(* Logix 5000 project; controller MV vendor 1 type 14 code 217 rev 31.11; software revision 31.00; part 14 of 53 *)
(* tags used below, declared in another part *)
   CWD : CHECKWORD_FLAGS;
   MC_copy_how_many : DINT;
   MC_data_file_value_to_move : DINT;
   MC_Delphi_I : DINT[60];
   MC_from_data_file : DINT;
   MC_from_data_offset : DINT;
   MC_LTX_001_1 : PlantItem;   // LTX_001_1
   MC_LTX_001_2 : PlantItem;   // LTX_001_2
   MC_LTX_001_3 : PlantItem;   // LTX_001_3
   MC_LTX_002_1 : PlantItem;   // LTX_002_1
   MC_LTX_002_2 : PlantItem;   // LTX_002_2
   MC_LTX_002_3 : PlantItem;   // LTX_002_3
   MC_LTX_003_1 : PlantItem;   // LTX_003_1
   MC_LTX_003_2 : PlantItem;   // LTX_003_2
   MC_LTX_003_3 : PlantItem;   // LTX_003_3
   MC_N10 : INT[255];   // SETTINGS
   MC_N100 : INT[255];   // C1_PLC Channel 1 PLC data
   MC_N101 : INT[255];   // CH1 PC>PLC Channel 1 PC to PLC
   MC_N102 : INT[255];   // CH1 PROG Channel 1 CIP progra m
   MC_N103 : INT[255];   // CH1 ITEMS Chwd.nos.of items to be checked for Chan nel 1
   MC_N104 : INT[255];   // CH1 REPORT Channel 1 CIP report file
   MC_N108 : INT[255];   // CH1 VDATA Channel 1 CIP progra m validation data
   MC_N112 : INT[255];   // FVR DATA Data read from FV ro uting PLC
   MC_N113 : INT[255];   // MVR DATA Data read from MV ro uting PLC
   MC_N114 : INT[255];   // YP DATA
   MC_N120 : INT[255];   // C2 PLC Channel 2 PLC data
   MC_N121 : INT[255];   // CH2 PC>PLC Channel 2 PC to PLC
   MC_N122 : INT[255];   // CH2 PROG Channel 2 CIP progra m
   MC_N123 : INT[255];   // CH2 ITEMS Chwd.nos.of items to be checked for Chan nel 2
   MC_N124 : INT[255];   // CH2 REPORT Channel 2 CIP report file
   MC_N128 : INT[255];   // CH2 VDATA Channel 2 CIP progra m validation data
   MC_N160 : INT[255];   // P40 CHECK
   MC_N161 : INT[255];   // P41 CHECK
   MC_N162 : INT[255];   // P42 CHECK
   MC_N163 : INT[255];   // P43 CHECK
   MC_N164 : INT[255];   // P44 CHECK
   MC_N165 : INT[255];   // P45 CHECK
   MC_N166 : INT[255];   // P46 CHECK
   MC_N167 : INT[255];   // Original N File From SLC, No Description Available
   MC_N20 : INT[255];   // P1 PRESS Control block and da ta for P1 pressure P ID loop
   MC_N200 : INT[255];   // CHK_WORK Plant item fault che cking work area
   MC_N201 : INT[255];   // P1 CHECK CIP program 1 plant item check list
   MC_N202 : INT[255];   // P2 CHECK CIP program 2 plant item check list
   MC_N203 : INT[255];   // P3 CHECK CIP program 3 plant item check list
   MC_N204 : INT[255];   // P4 CHECK CIP program 4 plant item check list
   MC_N205 : INT[255];   // P5 CHECK CIP program 5 plant item check list
   MC_N206 : INT[255];   // P6 CHECK CIP program 6 plant item check list
   MC_N207 : INT[255];   // P7 CHECK CIP program 7 plant item check list
   MC_N208 : INT[255];   // P8 CHECK CIP program 8 plant item check list
   MC_N209 : INT[255];   // P9 CHECK CIP program 9 plant item check list
   MC_N21 : INT[255];   // P1 FLOW Control block and da ta for P1 flowrate P ID loop
   MC_N210 : INT[255];   // P10 CHECK CIP program 10 plant item check list
   MC_N211 : INT[255];   // P11 CHECK CIP program 11 plant item check list
   MC_N212 : INT[255];   // P12 CHECK CIP program 12 plant item check list
   MC_N213 : INT[255];   // P13 CHECK CIP program 13 plant item check list
   MC_N214 : INT[255];   // P14 CHECK CIP program 14 plant item check list
   MC_N215 : INT[255];   // P15 CHECK CIP program 15 plant item check list
   MC_N216 : INT[255];   // P16 CHECK CIP program 16 plant item check list
   MC_N217 : INT[255];   // P17 CHECK CIP program 17 plant item check list
   MC_N218 : INT[255];   // P18 CHECK CIP program 18 plant item check list
   MC_N219 : INT[255];   // P19 CHECK CIP program 19 plant item check list
   MC_N22 : INT[255];   // P2 PRESS Control block and da ta for P2 pressure P ID loop
   MC_N220 : INT[255];   // P20 CHECK CIP program 20 plant item check list
   MC_N221 : INT[255];   // P21 CHECK CIP program 21 plant item check list
   MC_N222 : INT[255];   // P22 CHECK CIP program 22 plant item check list
   MC_N223 : INT[255];   // P23 CHECK CIP program 23 plant item check list
   MC_N224 : INT[255];   // P24 CHECK CIP program 24 plant item check list
   MC_N225 : INT[255];   // P25 CHECK CIP program 25 plant item check list
   MC_N226 : INT[255];   // P26 CHECK CIP program 26 plant item check list
   MC_N227 : INT[255];   // P27 CHECK CIP program 27 plant item check list
   MC_N228 : INT[255];   // P28 CHECK CIP program 28 plant item check list
   MC_N229 : INT[255];   // P29 CHECK CIP program 29 plant item check list
   MC_N23 : INT[255];   // P2 FLOW Control block and da ta for P2 flowrate P ID loop
   MC_N230 : INT[255];   // P30 CHECK CIP program 30 plant item check list
   MC_N231 : INT[255];   // P31 CHECK CIP program 31 plant item check list
   MC_N232 : INT[255];   // P32 CHECK CIP program 32 plant item check list
   MC_N233 : INT[255];   // P33 CHECK CIP program 33 plant item check list
   MC_N234 : INT[255];   // P34 CHECK CIP program 34 plant item check list
   MC_N235 : INT[255];   // P35 CHECK CIP program 35 plant item check list
   MC_N236 : INT[255];   // P36 CHECK CIP program 36 plant item check list
   MC_N237 : INT[255];   // P37 CHECK CIP program 37 plant item check list
   MC_N238 : INT[255];   // P38 CHECK CIP program 38 plant item check list
   MC_N239 : INT[255];   // P39 CHECK CIP program 39 plant item check list
   MC_N245 : INT[255];   // CC_WORK Continuous checking program work area
   MC_N7 : INT[255];   // INTEGER
   MC_N80 : INT[255];   // SRV1_PLC Detergent tank 1 ser vice PLC data
   MC_N81 : INT[255];   // SV1_PC Detergent tank 1 ser vice PC to PLC data
   MC_N82 : INT[255];   // SV1 ITEMS Chwd.nos.of items to be checked for DT1 service
   MC_N90 : INT[255];   // SV2_PLC Detergent tank 2 ser vice PLC data
   MC_N91 : INT[255];   // SV2_PC Detergent tank 2 ser vice PC to PLC data
   MC_N92 : INT[255];   // SV2 ITEMS Chwd.nos.of items to be checked for DT2 service
   MC_PX_100 : PlantItem;   // PX_100
   MC_PX_100_RawInput : ALIAS FOR RIO_Rack_2:11:I.Data.18;   // MC_PX_100
   MC_PX_101 : PlantItem;   // PX_101
   MC_PX_101_RawInput : ALIAS FOR RIO_Rack_2:11:I.Data.19;   // MC_PX_101
   MC_R2_SW1 : PlantItem;   // R2_SW1
   MC_R2_SW1_RawInput : ALIAS FOR RIO_Rack_2:12:I.Data.0;   // MC_R2_SW1
   MC_R2_SW2 : PlantItem;   // R2_SW2
   MC_R2_SW2_RawInput : ALIAS FOR RIO_Rack_2:12:I.Data.1;   // MC_R2_SW2
   MC_R2_SW3 : PlantItem;   // R2_SW3
   MC_R2_SW3_1 : PlantItem;   // R2_SW3_1
   MC_R2_SW3_1_RawInput : ALIAS FOR RIO_Rack_2:12:I.Data.3;   // MC_R2_SW3_1
   MC_R2_SW3_RawInput : ALIAS FOR RIO_Rack_2:12:I.Data.2;   // MC_R2_SW3
   MC_R2_SW4 : PlantItem;   // R2_SW4
   MC_R2_SW4_RawInput : ALIAS FOR RIO_Rack_2:12:I.Data.4;   // MC_R2_SW4
   MC_R3_SW1 : PlantItem;   // R3_SW1
   MC_R3_SW1_RawInput : ALIAS FOR RIO_Rack_2:12:I.Data.5;   // MC_R3_SW1
   MC_R3_SW2 : PlantItem;   // R3_SW2
   MC_R3_SW2_RawInput : ALIAS FOR RIO_Rack_2:12:I.Data.6;   // MC_R3_SW2
   MC_T4 : TIMER[255];   // TIMER
   MC_to_data_file : DINT;
   MC_to_data_offset : DINT;
   One_Second_One_Scan : ALIAS FOR One_Second_1_scan;
(* MC_Common, continued *)

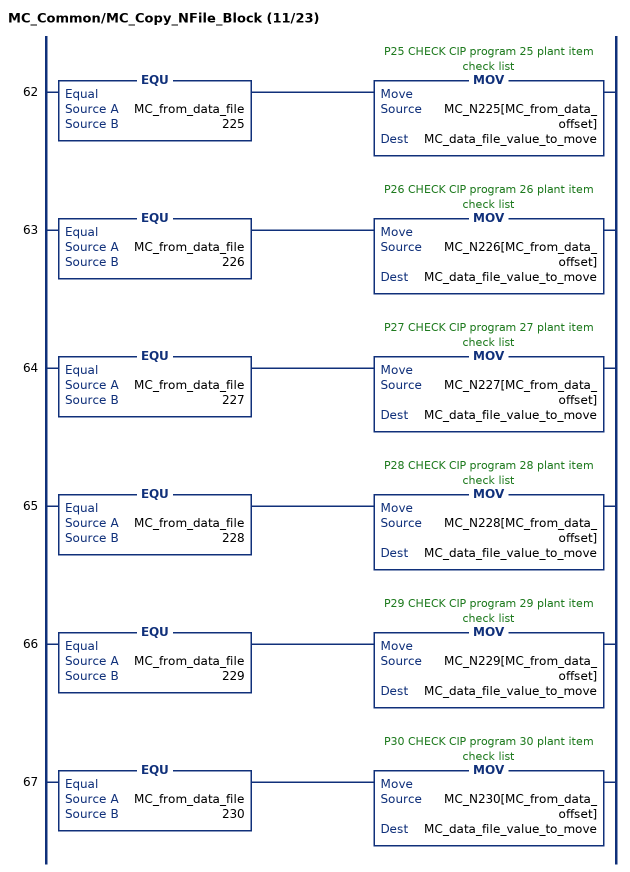
   [picture p203: MC_Common/MC_Copy_NFile_Block rungs 62-67]
   62: EQU(MC_from_data_file,225)MOV(MC_N225[MC_from_data_offset],MC_data_file_value_to_move);
   63: EQU(MC_from_data_file,226)MOV(MC_N226[MC_from_data_offset],MC_data_file_value_to_move);
   64: EQU(MC_from_data_file,227)MOV(MC_N227[MC_from_data_offset],MC_data_file_value_to_move);
   65: EQU(MC_from_data_file,228)MOV(MC_N228[MC_from_data_offset],MC_data_file_value_to_move);
   66: EQU(MC_from_data_file,229)MOV(MC_N229[MC_from_data_offset],MC_data_file_value_to_move);
   67: EQU(MC_from_data_file,230)MOV(MC_N230[MC_from_data_offset],MC_data_file_value_to_move);
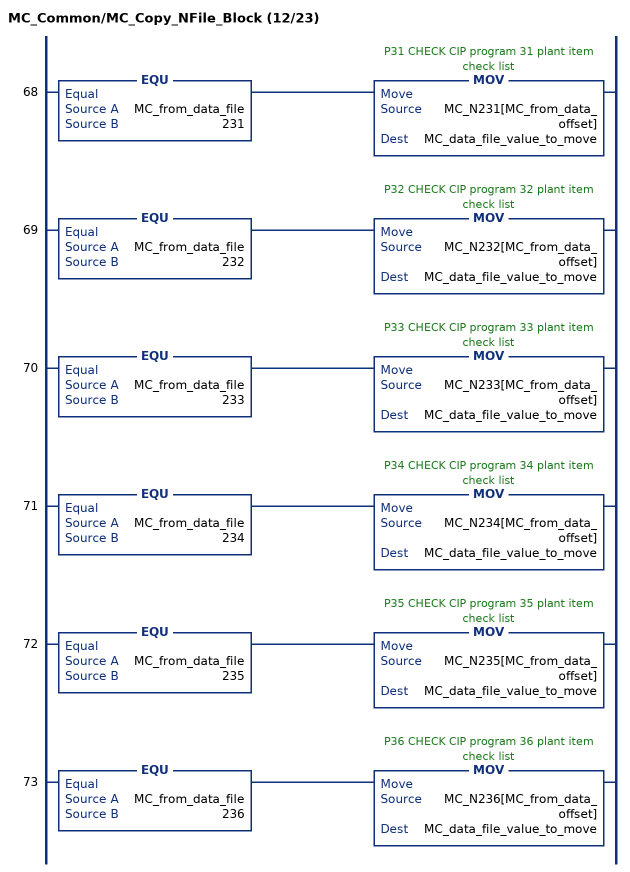
   68: EQU(MC_from_data_file,231)MOV(MC_N231[MC_from_data_offset],MC_data_file_value_to_move);
   69: EQU(MC_from_data_file,232)MOV(MC_N232[MC_from_data_offset],MC_data_file_value_to_move);
   70: EQU(MC_from_data_file,233)MOV(MC_N233[MC_from_data_offset],MC_data_file_value_to_move);
   71: EQU(MC_from_data_file,234)MOV(MC_N234[MC_from_data_offset],MC_data_file_value_to_move);
   72: EQU(MC_from_data_file,235)MOV(MC_N235[MC_from_data_offset],MC_data_file_value_to_move);
   73: EQU(MC_from_data_file,236)MOV(MC_N236[MC_from_data_offset],MC_data_file_value_to_move);
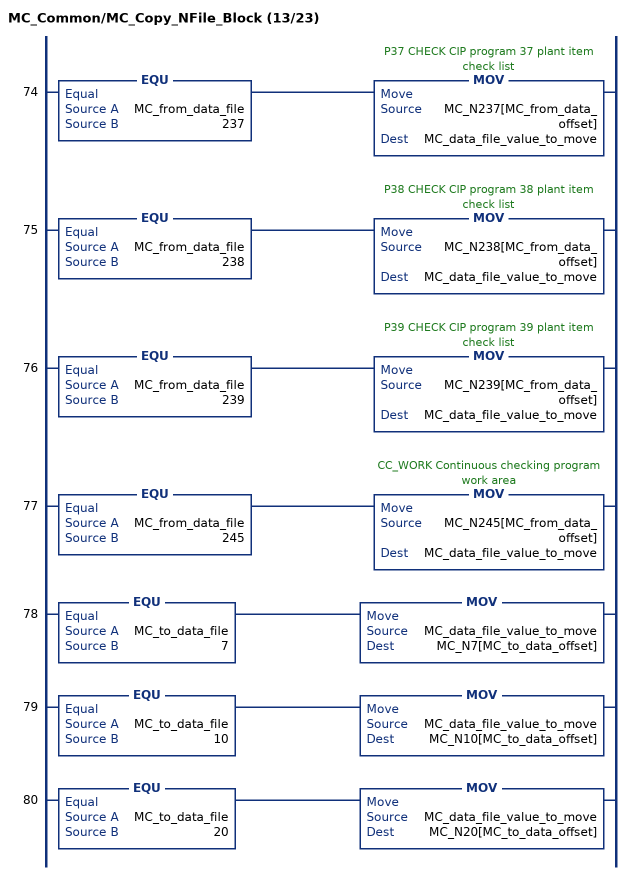
   74: EQU(MC_from_data_file,237)MOV(MC_N237[MC_from_data_offset],MC_data_file_value_to_move);
   75: EQU(MC_from_data_file,238)MOV(MC_N238[MC_from_data_offset],MC_data_file_value_to_move);
   76: EQU(MC_from_data_file,239)MOV(MC_N239[MC_from_data_offset],MC_data_file_value_to_move);
   77: EQU(MC_from_data_file,245)MOV(MC_N245[MC_from_data_offset],MC_data_file_value_to_move);
   78: EQU(MC_to_data_file,7)MOV(MC_data_file_value_to_move,MC_N7[MC_to_data_offset]);
   79: EQU(MC_to_data_file,10)MOV(MC_data_file_value_to_move,MC_N10[MC_to_data_offset]);
   80: EQU(MC_to_data_file,20)MOV(MC_data_file_value_to_move,MC_N20[MC_to_data_offset]);
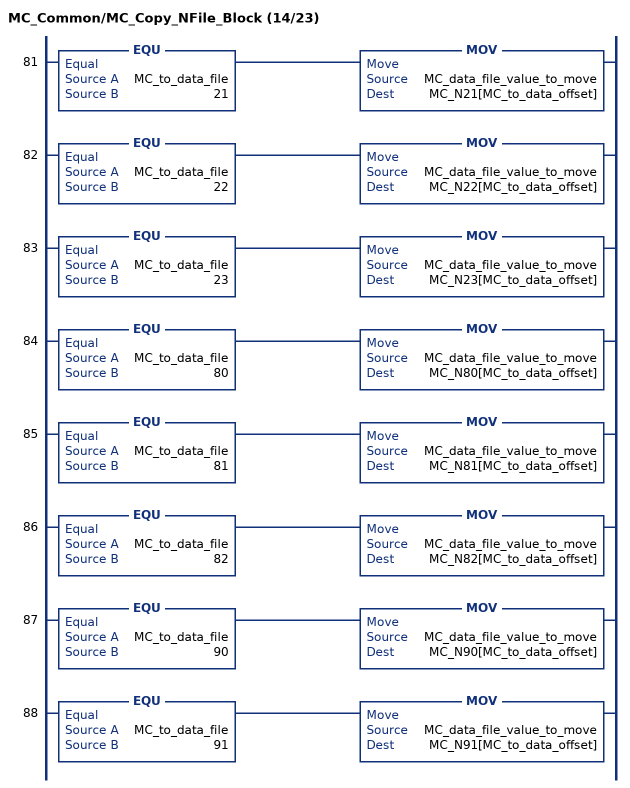
   81: EQU(MC_to_data_file,21)MOV(MC_data_file_value_to_move,MC_N21[MC_to_data_offset]);
   82: EQU(MC_to_data_file,22)MOV(MC_data_file_value_to_move,MC_N22[MC_to_data_offset]);
   83: EQU(MC_to_data_file,23)MOV(MC_data_file_value_to_move,MC_N23[MC_to_data_offset]);
   84: EQU(MC_to_data_file,80)MOV(MC_data_file_value_to_move,MC_N80[MC_to_data_offset]);
   85: EQU(MC_to_data_file,81)MOV(MC_data_file_value_to_move,MC_N81[MC_to_data_offset]);
   86: EQU(MC_to_data_file,82)MOV(MC_data_file_value_to_move,MC_N82[MC_to_data_offset]);
   87: EQU(MC_to_data_file,90)MOV(MC_data_file_value_to_move,MC_N90[MC_to_data_offset]);
   88: EQU(MC_to_data_file,91)MOV(MC_data_file_value_to_move,MC_N91[MC_to_data_offset]);
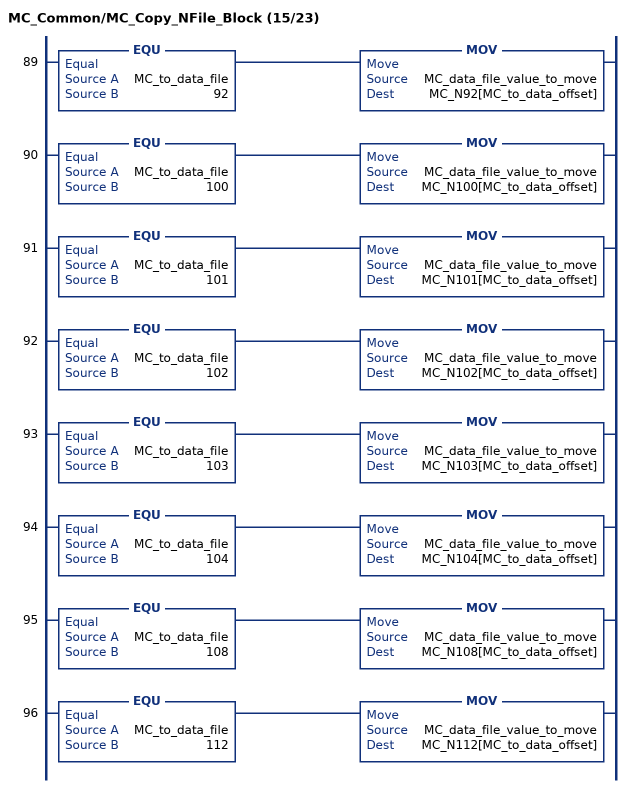
   89: EQU(MC_to_data_file,92)MOV(MC_data_file_value_to_move,MC_N92[MC_to_data_offset]);
   90: EQU(MC_to_data_file,100)MOV(MC_data_file_value_to_move,MC_N100[MC_to_data_offset]);
   91: EQU(MC_to_data_file,101)MOV(MC_data_file_value_to_move,MC_N101[MC_to_data_offset]);
   92: EQU(MC_to_data_file,102)MOV(MC_data_file_value_to_move,MC_N102[MC_to_data_offset]);
   93: EQU(MC_to_data_file,103)MOV(MC_data_file_value_to_move,MC_N103[MC_to_data_offset]);
   94: EQU(MC_to_data_file,104)MOV(MC_data_file_value_to_move,MC_N104[MC_to_data_offset]);
   95: EQU(MC_to_data_file,108)MOV(MC_data_file_value_to_move,MC_N108[MC_to_data_offset]);
   96: EQU(MC_to_data_file,112)MOV(MC_data_file_value_to_move,MC_N112[MC_to_data_offset]);
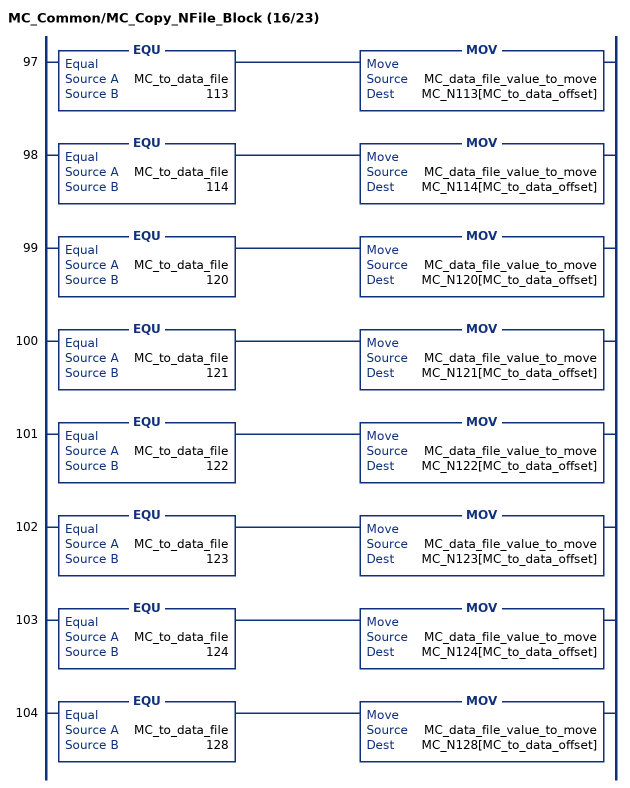
   97: EQU(MC_to_data_file,113)MOV(MC_data_file_value_to_move,MC_N113[MC_to_data_offset]);
   98: EQU(MC_to_data_file,114)MOV(MC_data_file_value_to_move,MC_N114[MC_to_data_offset]);
   99: EQU(MC_to_data_file,120)MOV(MC_data_file_value_to_move,MC_N120[MC_to_data_offset]);
   100: EQU(MC_to_data_file,121)MOV(MC_data_file_value_to_move,MC_N121[MC_to_data_offset]);
   101: EQU(MC_to_data_file,122)MOV(MC_data_file_value_to_move,MC_N122[MC_to_data_offset]);
   102: EQU(MC_to_data_file,123)MOV(MC_data_file_value_to_move,MC_N123[MC_to_data_offset]);
   103: EQU(MC_to_data_file,124)MOV(MC_data_file_value_to_move,MC_N124[MC_to_data_offset]);
   104: EQU(MC_to_data_file,128)MOV(MC_data_file_value_to_move,MC_N128[MC_to_data_offset]);
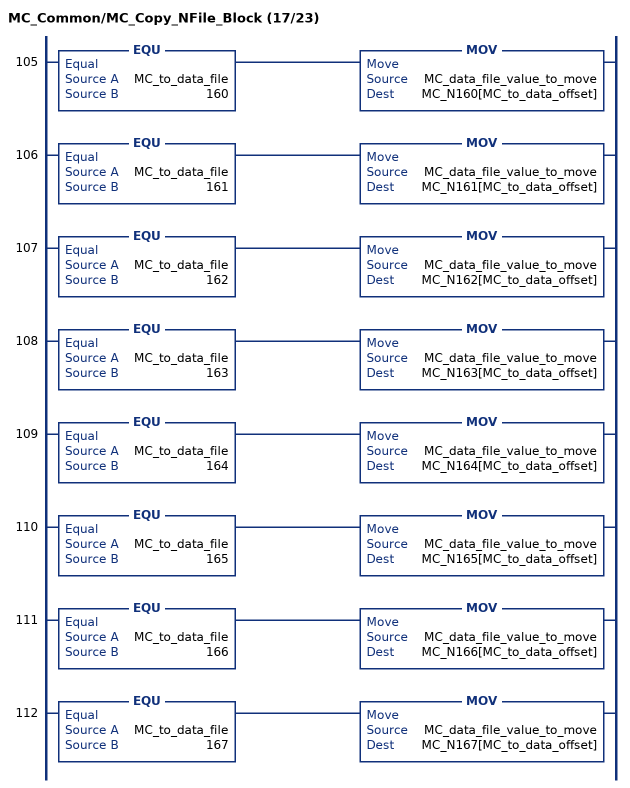
   105: EQU(MC_to_data_file,160)MOV(MC_data_file_value_to_move,MC_N160[MC_to_data_offset]);
   106: EQU(MC_to_data_file,161)MOV(MC_data_file_value_to_move,MC_N161[MC_to_data_offset]);
   107: EQU(MC_to_data_file,162)MOV(MC_data_file_value_to_move,MC_N162[MC_to_data_offset]);
   108: EQU(MC_to_data_file,163)MOV(MC_data_file_value_to_move,MC_N163[MC_to_data_offset]);
   109: EQU(MC_to_data_file,164)MOV(MC_data_file_value_to_move,MC_N164[MC_to_data_offset]);
   110: EQU(MC_to_data_file,165)MOV(MC_data_file_value_to_move,MC_N165[MC_to_data_offset]);
   111: EQU(MC_to_data_file,166)MOV(MC_data_file_value_to_move,MC_N166[MC_to_data_offset]);
   112: EQU(MC_to_data_file,167)MOV(MC_data_file_value_to_move,MC_N167[MC_to_data_offset]);
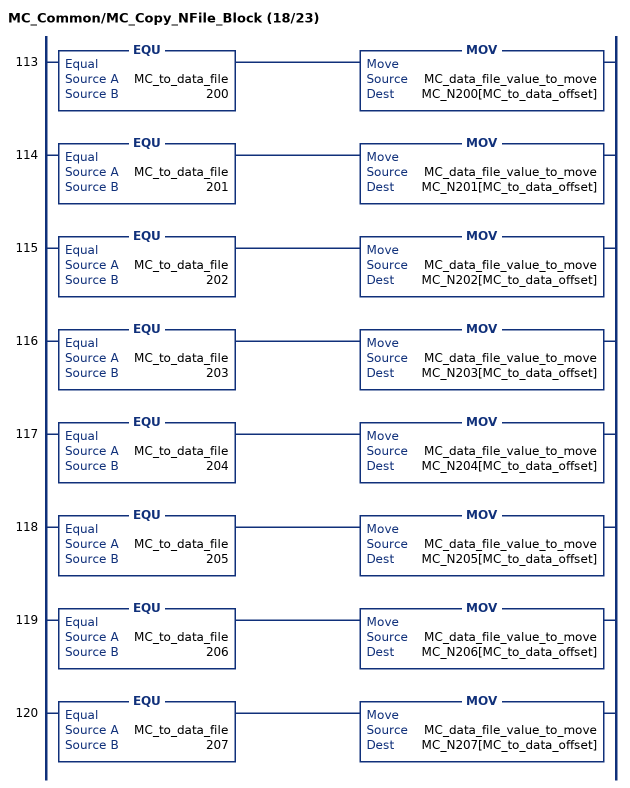
   113: EQU(MC_to_data_file,200)MOV(MC_data_file_value_to_move,MC_N200[MC_to_data_offset]);
   114: EQU(MC_to_data_file,201)MOV(MC_data_file_value_to_move,MC_N201[MC_to_data_offset]);
   115: EQU(MC_to_data_file,202)MOV(MC_data_file_value_to_move,MC_N202[MC_to_data_offset]);
   116: EQU(MC_to_data_file,203)MOV(MC_data_file_value_to_move,MC_N203[MC_to_data_offset]);
   117: EQU(MC_to_data_file,204)MOV(MC_data_file_value_to_move,MC_N204[MC_to_data_offset]);
   118: EQU(MC_to_data_file,205)MOV(MC_data_file_value_to_move,MC_N205[MC_to_data_offset]);
   119: EQU(MC_to_data_file,206)MOV(MC_data_file_value_to_move,MC_N206[MC_to_data_offset]);
   120: EQU(MC_to_data_file,207)MOV(MC_data_file_value_to_move,MC_N207[MC_to_data_offset]);
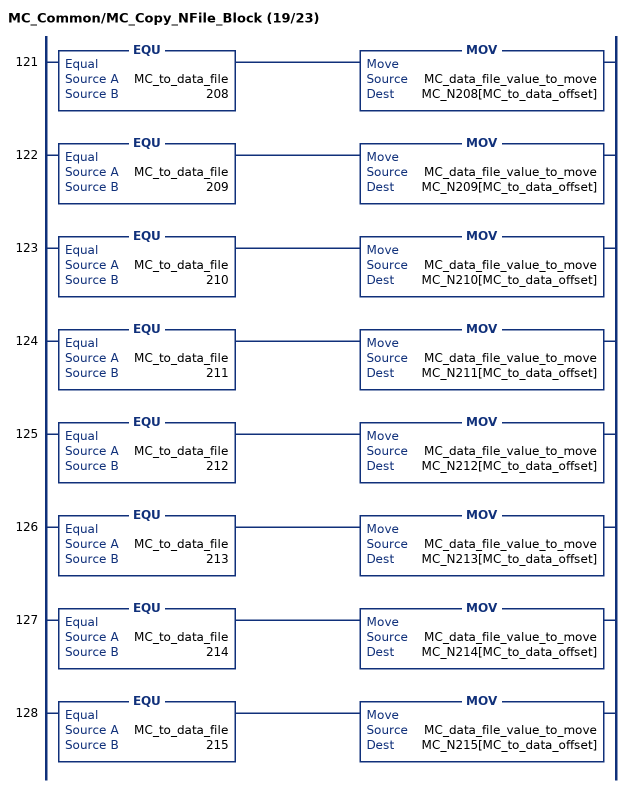
   121: EQU(MC_to_data_file,208)MOV(MC_data_file_value_to_move,MC_N208[MC_to_data_offset]);
   122: EQU(MC_to_data_file,209)MOV(MC_data_file_value_to_move,MC_N209[MC_to_data_offset]);
   123: EQU(MC_to_data_file,210)MOV(MC_data_file_value_to_move,MC_N210[MC_to_data_offset]);
   124: EQU(MC_to_data_file,211)MOV(MC_data_file_value_to_move,MC_N211[MC_to_data_offset]);
   125: EQU(MC_to_data_file,212)MOV(MC_data_file_value_to_move,MC_N212[MC_to_data_offset]);
   126: EQU(MC_to_data_file,213)MOV(MC_data_file_value_to_move,MC_N213[MC_to_data_offset]);
   127: EQU(MC_to_data_file,214)MOV(MC_data_file_value_to_move,MC_N214[MC_to_data_offset]);
   128: EQU(MC_to_data_file,215)MOV(MC_data_file_value_to_move,MC_N215[MC_to_data_offset]);
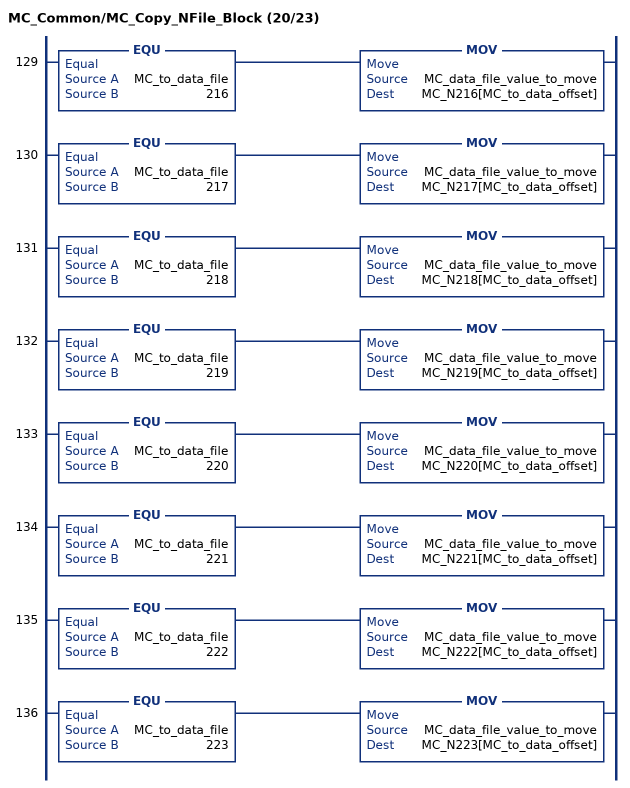
   129: EQU(MC_to_data_file,216)MOV(MC_data_file_value_to_move,MC_N216[MC_to_data_offset]);
   130: EQU(MC_to_data_file,217)MOV(MC_data_file_value_to_move,MC_N217[MC_to_data_offset]);
   131: EQU(MC_to_data_file,218)MOV(MC_data_file_value_to_move,MC_N218[MC_to_data_offset]);
   132: EQU(MC_to_data_file,219)MOV(MC_data_file_value_to_move,MC_N219[MC_to_data_offset]);
   133: EQU(MC_to_data_file,220)MOV(MC_data_file_value_to_move,MC_N220[MC_to_data_offset]);
   134: EQU(MC_to_data_file,221)MOV(MC_data_file_value_to_move,MC_N221[MC_to_data_offset]);
   135: EQU(MC_to_data_file,222)MOV(MC_data_file_value_to_move,MC_N222[MC_to_data_offset]);
   136: EQU(MC_to_data_file,223)MOV(MC_data_file_value_to_move,MC_N223[MC_to_data_offset]);
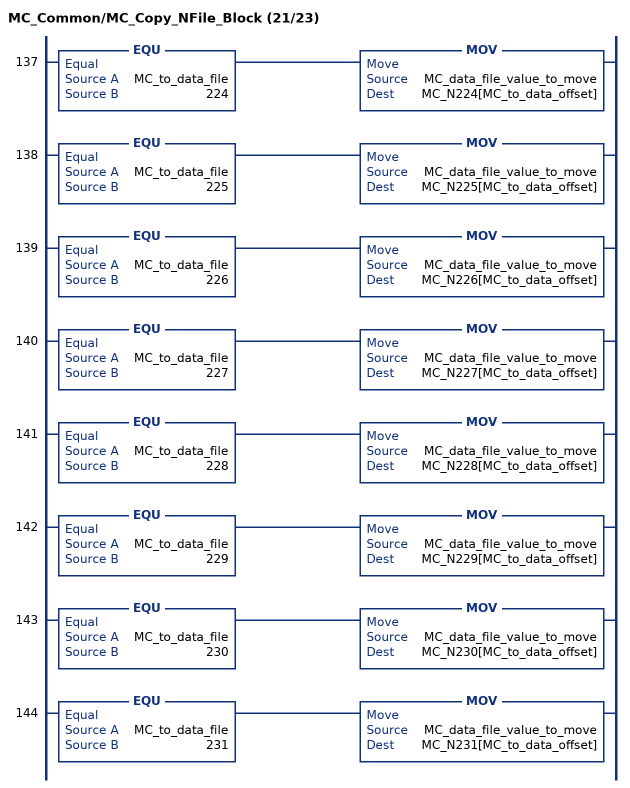
   137: EQU(MC_to_data_file,224)MOV(MC_data_file_value_to_move,MC_N224[MC_to_data_offset]);
   138: EQU(MC_to_data_file,225)MOV(MC_data_file_value_to_move,MC_N225[MC_to_data_offset]);
   139: EQU(MC_to_data_file,226)MOV(MC_data_file_value_to_move,MC_N226[MC_to_data_offset]);
   140: EQU(MC_to_data_file,227)MOV(MC_data_file_value_to_move,MC_N227[MC_to_data_offset]);
   141: EQU(MC_to_data_file,228)MOV(MC_data_file_value_to_move,MC_N228[MC_to_data_offset]);
   142: EQU(MC_to_data_file,229)MOV(MC_data_file_value_to_move,MC_N229[MC_to_data_offset]);
   143: EQU(MC_to_data_file,230)MOV(MC_data_file_value_to_move,MC_N230[MC_to_data_offset]);
   144: EQU(MC_to_data_file,231)MOV(MC_data_file_value_to_move,MC_N231[MC_to_data_offset]);
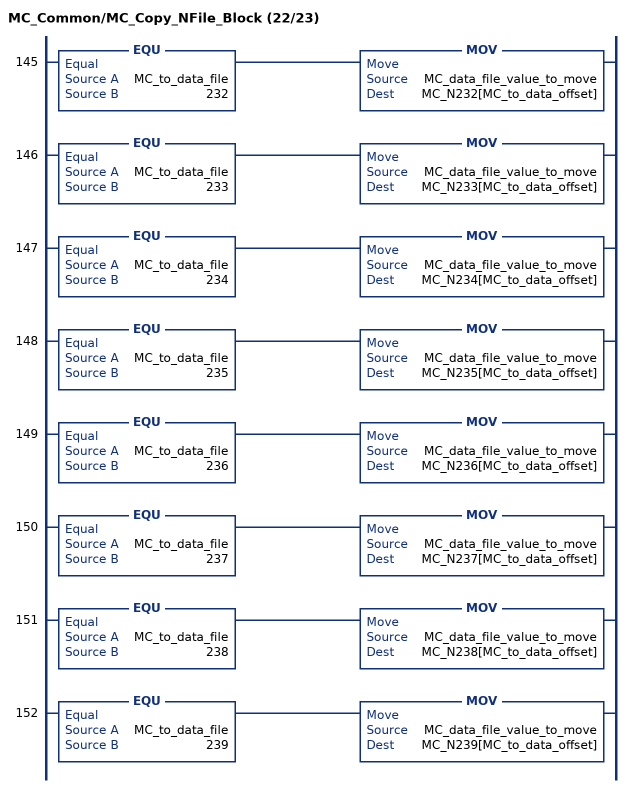
   145: EQU(MC_to_data_file,232)MOV(MC_data_file_value_to_move,MC_N232[MC_to_data_offset]);
   146: EQU(MC_to_data_file,233)MOV(MC_data_file_value_to_move,MC_N233[MC_to_data_offset]);
   147: EQU(MC_to_data_file,234)MOV(MC_data_file_value_to_move,MC_N234[MC_to_data_offset]);
   148: EQU(MC_to_data_file,235)MOV(MC_data_file_value_to_move,MC_N235[MC_to_data_offset]);
   149: EQU(MC_to_data_file,236)MOV(MC_data_file_value_to_move,MC_N236[MC_to_data_offset]);
   150: EQU(MC_to_data_file,237)MOV(MC_data_file_value_to_move,MC_N237[MC_to_data_offset]);
   151: EQU(MC_to_data_file,238)MOV(MC_data_file_value_to_move,MC_N238[MC_to_data_offset]);
   152: EQU(MC_to_data_file,239)MOV(MC_data_file_value_to_move,MC_N239[MC_to_data_offset]);